HMI tags "Process_Value"
   "DB602_PV_Tank_Tank{0}_Temp_PV_Conf_ActV_ModulNo" : Int = PLC DB602_PV_Tank.Tank[0].Temp.PV_Conf_ActV.ModulNo AT %DB602.DBW32, 1 s
      on ChangeValue: SetBit("DB702_Tank_Value.Write")
   "DB602_PV_Tank_Tank{0}_Temp_PV_Conf_ActV_Address" : Int = PLC DB602_PV_Tank.Tank[0].Temp.PV_Conf_ActV.Address AT %DB602.DBW34, 1 s
      on ChangeValue: SetBit("DB702_Tank_Value.Write")
   "DB602_PV_Tank_Tank{0}_Temp_PV_Conf_ActV_OffsetSignal" : Int = PLC DB602_PV_Tank.Tank[0].Temp.PV_Conf_ActV.OffsetSignal AT %DB602.DBW36, 1 s
      on ChangeValue: SetBit("DB702_Tank_Value.Write")
   "DB602_PV_Tank_Tank{0}_Temp_PV_Conf_ActV_Multiplier" : Real = PLC DB602_PV_Tank.Tank[0].Temp.PV_Conf_ActV.Multiplier AT %DB602.DBD38, 1 s
      on ChangeValue: SetBit("DB702_Tank_Value.Write")
   "DB602_PV_Tank_Tank{0}_Temp_PV_Conf_ActV_MinValueSensor" : Real = PLC DB602_PV_Tank.Tank[0].Temp.PV_Conf_ActV.MinValueSensor AT %DB602.DBD42, 1 s
      on ChangeValue: SetBit("DB702_Tank_Value.Write")
   "DB602_PV_Tank_Tank{0}_Temp_PV_Conf_ActV_MaxValueSensor" : Real = PLC DB602_PV_Tank.Tank[0].Temp.PV_Conf_ActV.MaxValueSensor AT %DB602.DBD46, 1 s
      on ChangeValue: SetBit("DB702_Tank_Value.Write")
   "DB602_PV_Tank_Tank{0}_Temp_PV_Conf_ActV_MaxSignalResolution" : Real = PLC DB602_PV_Tank.Tank[0].Temp.PV_Conf_ActV.MaxSignalResolution AT %DB602.DBD50, 1 s
      on ChangeValue: SetBit("DB702_Tank_Value.Write")
   "DB602_PV_Tank_Tank{0}_Temp_PV_ActV_Value" : Real = PLC DB602_PV_Tank.Tank[0].Temp.PV_ActV.Value AT %DB602.DBD26, 1 s
      on ChangeValue: SetBit("DB702_Tank_Value.Write")
   "DB602_PV_Tank_Tank{0}_Level_PV_ActV_Value" : Real = PLC DB602_PV_Tank.Tank[0].Level.PV_ActV.Value AT %DB602.DBD74, 1 s
      on ChangeValue: SetBit("DB702_Tank_Value.Write")
   "DB602_PV_Tank_Tank{0}_Level_PV_Conf_ActV_ModulNo" : Int = PLC DB602_PV_Tank.Tank[0].Level.PV_Conf_ActV.ModulNo AT %DB602.DBW80, 1 s
      on ChangeValue: SetBit("DB702_Tank_Value.Write")
   "DB602_PV_Tank_Tank{0}_Level_PV_Conf_ActV_Address" : Int = PLC DB602_PV_Tank.Tank[0].Level.PV_Conf_ActV.Address AT %DB602.DBW82, 1 s
      on ChangeValue: SetBit("DB702_Tank_Value.Write")
   "DB602_PV_Tank_Tank{0}_Level_PV_Conf_ActV_OffsetSignal" : Int = PLC DB602_PV_Tank.Tank[0].Level.PV_Conf_ActV.OffsetSignal AT %DB602.DBW84, 1 s
      on ChangeValue: SetBit("DB702_Tank_Value.Write")
   "DB602_PV_Tank_Tank{0}_Level_PV_Conf_ActV_Multiplier" : Real = PLC DB602_PV_Tank.Tank[0].Level.PV_Conf_ActV.Multiplier AT %DB602.DBD86, 1 s
      on ChangeValue: SetBit("DB702_Tank_Value.Write")
   "DB602_PV_Tank_Tank{0}_Level_PV_Conf_ActV_MinValueSensor" : Real = PLC DB602_PV_Tank.Tank[0].Level.PV_Conf_ActV.MinValueSensor AT %DB602.DBD90, 1 s
      on ChangeValue: SetBit("DB702_Tank_Value.Write")
   "DB602_PV_Tank_Tank{0}_Level_PV_Conf_ActV_MaxValueSensor" : Real = PLC DB602_PV_Tank.Tank[0].Level.PV_Conf_ActV.MaxValueSensor AT %DB602.DBD94, 1 s
      on ChangeValue: SetBit("DB702_Tank_Value.Write")
   "DB602_PV_Tank_Tank{0}_Level_PV_Conf_ActV_MaxSignalResolution" : Real = PLC DB602_PV_Tank.Tank[0].Level.PV_Conf_ActV.MaxSignalResolution AT %DB602.DBD98, 1 s
      on ChangeValue: SetBit("DB702_Tank_Value.Write")
   "DB602_PV_Tank_Tank{0}_Nucleation_PV_Conf_ActV_ModulNo" : Int = PLC DB602_PV_Tank.Tank[0].Nucleation.PV_Conf_ActV.ModulNo AT %DB602.DBW176, 1 s
      on ChangeValue: SetBit("DB702_Tank_Value.Write")
   "DB602_PV_Tank_Tank{0}_Nucleation_PV_Conf_ActV_Address" : Int = PLC DB602_PV_Tank.Tank[0].Nucleation.PV_Conf_ActV.Address AT %DB602.DBW178, 1 s
      on ChangeValue: SetBit("DB702_Tank_Value.Write")
   "DB602_PV_Tank_Tank{0}_Nucleation_PV_Conf_ActV_OffsetSignal" : Int = PLC DB602_PV_Tank.Tank[0].Nucleation.PV_Conf_ActV.OffsetSignal AT %DB602.DBW180, 1 s
      on ChangeValue: SetBit("DB702_Tank_Value.Write")
   "DB602_PV_Tank_Tank{0}_Nucleation_PV_Conf_ActV_Multiplier" : Real = PLC DB602_PV_Tank.Tank[0].Nucleation.PV_Conf_ActV.Multiplier AT %DB602.DBD182, 1 s
      on ChangeValue: SetBit("DB702_Tank_Value.Write")
   "DB602_PV_Tank_Tank{0}_Nucleation_PV_Conf_ActV_MinValueSensor" : Real = PLC DB602_PV_Tank.Tank[0].Nucleation.PV_Conf_ActV.MinValueSensor AT %DB602.DBD186, 1 s
      on ChangeValue: SetBit("DB702_Tank_Value.Write")
   "DB602_PV_Tank_Tank{0}_Nucleation_PV_Conf_ActV_MaxValueSensor" : Real = PLC DB602_PV_Tank.Tank[0].Nucleation.PV_Conf_ActV.MaxValueSensor AT %DB602.DBD190, 1 s
      on ChangeValue: SetBit("DB702_Tank_Value.Write")
   "DB602_PV_Tank_Tank{0}_Nucleation_PV_Conf_ActV_MaxSignalResolution" : Real = PLC DB602_PV_Tank.Tank[0].Nucleation.PV_Conf_ActV.MaxSignalResolution AT %DB602.DBD194, 1 s
      on ChangeValue: SetBit("DB702_Tank_Value.Write")
   "DB602_PV_Tank_Tank{0}_Nucleation_PV_ActV_Value" : Real = PLC DB602_PV_Tank.Tank[0].Nucleation.PV_ActV.Value AT %DB602.DBD170, 1 s
      on ChangeValue: SetBit("DB702_Tank_Value.Write")
   "DB702_Tank_Value_Read" : Bool = PLC DB702_Tank_Value.Read AT %DB702.DBX4.0, 1 s
   "DB608_PV_Metering_Metering{0}_Flow_PV_Conf_ActV_Address" : Int = PLC DB608_PV_Metering.Metering[0].Flow.PV_Conf_ActV.Address AT %DB608.DBW34, 1 s
      on ChangeValue: SetBit("DB608_PV_Metering_Write")
   "DB608_PV_Metering_Metering{0}_Flow_PV_ActV_Value" : Real = PLC DB608_PV_Metering.Metering[0].Flow.PV_ActV.Value AT %DB608.DBD26, 1 s
      on ChangeValue: SetBit("DB608_PV_Metering_Write")
   "DB608_PV_Metering_Metering{0}_Pressure_PV_Conf_ActV_ModulNo" : Int = PLC DB608_PV_Metering.Metering[0].Pressure.PV_Conf_ActV.ModulNo AT %DB608.DBW80, 1 s
      on ChangeValue: SetBit("DB608_PV_Metering_Write")
   "DB608_PV_Metering_Metering{0}_Pressure_PV_Conf_ActV_Address" : Int = PLC DB608_PV_Metering.Metering[0].Pressure.PV_Conf_ActV.Address AT %DB608.DBW82, 1 s
      on ChangeValue: SetBit("DB608_PV_Metering_Write")
   "DB608_PV_Metering_Metering{0}_Pressure_PV_Conf_ActV_OffsetSignal" : Int = PLC DB608_PV_Metering.Metering[0].Pressure.PV_Conf_ActV.OffsetSignal AT %DB608.DBW84, 1 s
      on ChangeValue: SetBit("DB608_PV_Metering_Write")
   "DB608_PV_Metering_Metering{0}_Pressure_PV_Conf_ActV_Multiplier" : Real = PLC DB608_PV_Metering.Metering[0].Pressure.PV_Conf_ActV.Multiplier AT %DB608.DBD86, 1 s
      on ChangeValue: SetBit("DB608_PV_Metering_Write")
   "DB608_PV_Metering_Metering{0}_Pressure_PV_Conf_ActV_MinValueSensor" : Real = PLC DB608_PV_Metering.Metering[0].Pressure.PV_Conf_ActV.MinValueSensor AT %DB608.DBD90, 1 s
      on ChangeValue: SetBit("DB608_PV_Metering_Write")
   "DB608_PV_Metering_Metering{0}_Pressure_PV_Conf_ActV_MaxValueSensor" : Real = PLC DB608_PV_Metering.Metering[0].Pressure.PV_Conf_ActV.MaxValueSensor AT %DB608.DBD94, 1 s
      on ChangeValue: SetBit("DB608_PV_Metering_Write")
   "DB608_PV_Metering_Metering{0}_Pressure_PV_Conf_ActV_MaxSignalResolution" : Real = PLC DB608_PV_Metering.Metering[0].Pressure.PV_Conf_ActV.MaxSignalResolution AT %DB608.DBD98, 1 s
      on ChangeValue: SetBit("DB608_PV_Metering_Write")
   "DB608_PV_Metering_Metering{0}_Pressure_PV_ActV_Value" : Real = PLC DB608_PV_Metering.Metering[0].Pressure.PV_ActV.Value AT %DB608.DBD74, 1 s
      on ChangeValue: SetBit("DB608_PV_Metering_Write")
   "DB608_PV_Metering_Metering{0}_Temperature_PV_Conf_ActV_ModulNo" : Int = PLC DB608_PV_Metering.Metering[0].Temperature.PV_Conf_ActV.ModulNo AT %DB608.DBW128, 1 s
      on ChangeValue: SetBit("DB608_PV_Metering_Write")
   "DB608_PV_Metering_Metering{0}_Temperature_PV_Conf_ActV_Address" : Int = PLC DB608_PV_Metering.Metering[0].Temperature.PV_Conf_ActV.Address AT %DB608.DBW130, 1 s
      on ChangeValue: SetBit("DB608_PV_Metering_Write")
   "DB608_PV_Metering_Metering{0}_Temperature_PV_Conf_ActV_OffsetSignal" : Int = PLC DB608_PV_Metering.Metering[0].Temperature.PV_Conf_ActV.OffsetSignal AT %DB608.DBW132, 1 s
      on ChangeValue: SetBit("DB608_PV_Metering_Write")
   "DB608_PV_Metering_Metering{0}_Temperature_PV_Conf_ActV_Multiplier" : Real = PLC DB608_PV_Metering.Metering[0].Temperature.PV_Conf_ActV.Multiplier AT %DB608.DBD134, 1 s
      on ChangeValue: SetBit("DB608_PV_Metering_Write")
   "DB608_PV_Metering_Metering{0}_Temperature_PV_Conf_ActV_MinValueSensor" : Real = PLC DB608_PV_Metering.Metering[0].Temperature.PV_Conf_ActV.MinValueSensor AT %DB608.DBD138, 1 s
      on ChangeValue: SetBit("DB608_PV_Metering_Write")
   "DB608_PV_Metering_Metering{0}_Temperature_PV_Conf_ActV_MaxValueSensor" : Real = PLC DB608_PV_Metering.Metering[0].Temperature.PV_Conf_ActV.MaxValueSensor AT %DB608.DBD142, 1 s
      on ChangeValue: SetBit("DB608_PV_Metering_Write")
   "DB608_PV_Metering_Metering{0}_Temperature_PV_Conf_ActV_MaxSignalResolution" : Real = PLC DB608_PV_Metering.Metering[0].Temperature.PV_Conf_ActV.MaxSignalResolution AT %DB608.DBD146, 1 s
      on ChangeValue: SetBit("DB608_PV_Metering_Write")
   "DB608_PV_Metering_Metering{0}_Temperature_PV_ActV_Value" : Real = PLC DB608_PV_Metering.Metering[0].Temperature.PV_ActV.Value AT %DB608.DBD122, 1 s
      on ChangeValue: SetBit("DB608_PV_Metering_Write")
   "DB608_PV_Metering_Metering{0}_Pre_Pressure_PV_ActV_Value" : Real = PLC DB608_PV_Metering.Metering[0].Pre_Pressure.PV_ActV.Value AT %DB608.DBD170, 1 s
      on ChangeValue: SetBit("DB608_PV_Metering_Write")
   "DB608_PV_Metering_Metering{0}_Pre_Pressure_PV_Conf_ActV_ModulNo" : Int = PLC DB608_PV_Metering.Metering[0].Pre_Pressure.PV_Conf_ActV.ModulNo AT %DB608.DBW176, 1 s
      on ChangeValue: SetBit("DB608_PV_Metering_Write")
   "DB608_PV_Metering_Metering{0}_Pre_Pressure_PV_Conf_ActV_Address" : Int = PLC DB608_PV_Metering.Metering[0].Pre_Pressure.PV_Conf_ActV.Address AT %DB608.DBW178, 1 s
      on ChangeValue: SetBit("DB608_PV_Metering_Write")
   "DB608_PV_Metering_Metering{0}_Pre_Pressure_PV_Conf_ActV_OffsetSignal" : Int = PLC DB608_PV_Metering.Metering[0].Pre_Pressure.PV_Conf_ActV.OffsetSignal AT %DB608.DBW180, 1 s
      on ChangeValue: SetBit("DB608_PV_Metering_Write")
   "DB608_PV_Metering_Metering{0}_Pre_Pressure_PV_Conf_ActV_Multiplier" : Real = PLC DB608_PV_Metering.Metering[0].Pre_Pressure.PV_Conf_ActV.Multiplier AT %DB608.DBD182, 1 s
      on ChangeValue: SetBit("DB608_PV_Metering_Write")
   "DB608_PV_Metering_Metering{0}_Pre_Pressure_PV_Conf_ActV_MinValueSensor" : Real = PLC DB608_PV_Metering.Metering[0].Pre_Pressure.PV_Conf_ActV.MinValueSensor AT %DB608.DBD186, 1 s
      on ChangeValue: SetBit("DB608_PV_Metering_Write")
   "DB608_PV_Metering_Metering{0}_Pre_Pressure_PV_Conf_ActV_MaxValueSensor" : Real = PLC DB608_PV_Metering.Metering[0].Pre_Pressure.PV_Conf_ActV.MaxValueSensor AT %DB608.DBD190, 1 s
      on ChangeValue: SetBit("DB608_PV_Metering_Write")
   "DB608_PV_Metering_Metering{0}_Pre_Pressure_PV_Conf_ActV_MaxSignalResolution" : Real = PLC DB608_PV_Metering.Metering[0].Pre_Pressure.PV_Conf_ActV.MaxSignalResolution AT %DB608.DBD194, 1 s
      on ChangeValue: SetBit("DB608_PV_Metering_Write")
   "DB608_PV_Metering_HeatexchangerHP{0}_PV_ActV_Value" : Real = PLC DB608_PV_Metering.HeatexchangerHP[0].PV_ActV.Value AT %DB608.DBD3146, 1 s
      on ChangeValue: SetBit("DB608_PV_Metering_Write")
   "DB608_PV_Metering_HeatexchangerHP{0}_PV_Conf_ActV_ModulNo" : Int = PLC DB608_PV_Metering.HeatexchangerHP[0].PV_Conf_ActV.ModulNo AT %DB608.DBW3152, 1 s
      on ChangeValue: SetBit("DB608_PV_Metering_Write")
   "DB608_PV_Metering_HeatexchangerHP{0}_PV_Conf_ActV_Address" : Int = PLC DB608_PV_Metering.HeatexchangerHP[0].PV_Conf_ActV.Address AT %DB608.DBW3154, 1 s
      on ChangeValue: SetBit("DB608_PV_Metering_Write")
   "DB608_PV_Metering_HeatexchangerHP{0}_PV_Conf_ActV_OffsetSignal" : Int = PLC DB608_PV_Metering.HeatexchangerHP[0].PV_Conf_ActV.OffsetSignal AT %DB608.DBW3156, 1 s
      on ChangeValue: SetBit("DB608_PV_Metering_Write")
   "DB608_PV_Metering_HeatexchangerHP{0}_PV_Conf_ActV_Multiplier" : Real = PLC DB608_PV_Metering.HeatexchangerHP[0].PV_Conf_ActV.Multiplier AT %DB608.DBD3158, 1 s
      on ChangeValue: SetBit("DB608_PV_Metering_Write")
   "DB608_PV_Metering_HeatexchangerHP{0}_PV_Conf_ActV_MinValueSensor" : Real = PLC DB608_PV_Metering.HeatexchangerHP[0].PV_Conf_ActV.MinValueSensor AT %DB608.DBD3162, 1 s
      on ChangeValue: SetBit("DB608_PV_Metering_Write")
   "DB608_PV_Metering_HeatexchangerHP{0}_PV_Conf_ActV_MaxValueSensor" : Real = PLC DB608_PV_Metering.HeatexchangerHP[0].PV_Conf_ActV.MaxValueSensor AT %DB608.DBD3166, 1 s
      on ChangeValue: SetBit("DB608_PV_Metering_Write")
   "DB608_PV_Metering_HeatexchangerHP{0}_PV_Conf_ActV_MaxSignalResolution" : Real = PLC DB608_PV_Metering.HeatexchangerHP[0].PV_Conf_ActV.MaxSignalResolution AT %DB608.DBD3170, 1 s
      on ChangeValue: SetBit("DB608_PV_Metering_Write")
   "DB604_PV_Mixinghead_Mixinghead{0}_Inerting_PV_Conf_ActV_ModulNo" : Int = PLC DB604_PV_Mixinghead.Mixinghead[0].Inerting.PV_Conf_ActV.ModulNo AT %DB604.DBW704, 1 s
      on ChangeValue: SetBit("DB704_MH_Value_Write")
   "DB604_PV_Mixinghead_Mixinghead{0}_Inerting_PV_Conf_ActV_Address" : Int = PLC DB604_PV_Mixinghead.Mixinghead[0].Inerting.PV_Conf_ActV.Address AT %DB604.DBW706, 1 s
      on ChangeValue: SetBit("DB704_MH_Value_Write")
   "DB604_PV_Mixinghead_Mixinghead{0}_Inerting_PV_Conf_ActV_OffsetSignal" : Int = PLC DB604_PV_Mixinghead.Mixinghead[0].Inerting.PV_Conf_ActV.OffsetSignal AT %DB604.DBW708, 1 s
      on ChangeValue: SetBit("DB704_MH_Value_Write")
   "DB604_PV_Mixinghead_Mixinghead{0}_Inerting_PV_Conf_ActV_Multiplier" : Real = PLC DB604_PV_Mixinghead.Mixinghead[0].Inerting.PV_Conf_ActV.Multiplier AT %DB604.DBD710, 1 s
      on ChangeValue: SetBit("DB704_MH_Value_Write")
   "DB604_PV_Mixinghead_Mixinghead{0}_Inerting_PV_Conf_ActV_MinValueSensor" : Real = PLC DB604_PV_Mixinghead.Mixinghead[0].Inerting.PV_Conf_ActV.MinValueSensor AT %DB604.DBD714, 1 s
      on ChangeValue: SetBit("DB704_MH_Value_Write")
   "DB604_PV_Mixinghead_Mixinghead{0}_Inerting_PV_Conf_ActV_MaxValueSensor" : Real = PLC DB604_PV_Mixinghead.Mixinghead[0].Inerting.PV_Conf_ActV.MaxValueSensor AT %DB604.DBD718, 1 s
      on ChangeValue: SetBit("DB704_MH_Value_Write")
   "DB604_PV_Mixinghead_Mixinghead{0}_Inerting_PV_Conf_ActV_MaxSignalResolution" : Real = PLC DB604_PV_Mixinghead.Mixinghead[0].Inerting.PV_Conf_ActV.MaxSignalResolution AT %DB604.DBD722, 1 s
      on ChangeValue: SetBit("DB704_MH_Value_Write")
   "DB604_PV_Mixinghead_Mixinghead{0}_Inerting_PV_ActV_Value" : Real = PLC DB604_PV_Mixinghead.Mixinghead[0].Inerting.PV_ActV.Value AT %DB604.DBD698, 1 s
      on ChangeValue: SetBit("DB704_MH_Value_Write")
   "DB604_PV_Mixinghead_Mixinghead{0}_Pressure_Connection{1}_PV_Conf_ActV_ModulNo" : Int = PLC DB604_PV_Mixinghead.Mixinghead[0].Pressure_Connection[1].PV_Conf_ActV.ModulNo AT %DB604.DBW32, 1 s
      on ChangeValue: SetBit("DB704_MH_Value_Write")
   "DB604_PV_Mixinghead_Mixinghead{0}_Pressure_Connection{1}_PV_Conf_ActV_Address" : Int = PLC DB604_PV_Mixinghead.Mixinghead[0].Pressure_Connection[1].PV_Conf_ActV.Address AT %DB604.DBW34, 1 s
      on ChangeValue: SetBit("DB704_MH_Value_Write")
   "DB604_PV_Mixinghead_Mixinghead{0}_Pressure_Connection{1}_PV_Conf_ActV_OffsetSignal" : Int = PLC DB604_PV_Mixinghead.Mixinghead[0].Pressure_Connection[1].PV_Conf_ActV.OffsetSignal AT %DB604.DBW36, 1 s
      on ChangeValue: SetBit("DB704_MH_Value_Write")
   "DB604_PV_Mixinghead_Mixinghead{0}_Pressure_Connection{1}_PV_Conf_ActV_Multiplier" : Real = PLC DB604_PV_Mixinghead.Mixinghead[0].Pressure_Connection[1].PV_Conf_ActV.Multiplier AT %DB604.DBD38, 1 s
      on ChangeValue: SetBit("DB704_MH_Value_Write")
   "DB604_PV_Mixinghead_Mixinghead{0}_Pressure_Connection{1}_PV_Conf_ActV_MinValueSensor" : Real = PLC DB604_PV_Mixinghead.Mixinghead[0].Pressure_Connection[1].PV_Conf_ActV.MinValueSensor AT %DB604.DBD42, 1 s
      on ChangeValue: SetBit("DB704_MH_Value_Write")
   "DB604_PV_Mixinghead_Mixinghead{0}_Pressure_Connection{1}_PV_Conf_ActV_MaxValueSensor" : Real = PLC DB604_PV_Mixinghead.Mixinghead[0].Pressure_Connection[1].PV_Conf_ActV.MaxValueSensor AT %DB604.DBD46, 1 s
      on ChangeValue: SetBit("DB704_MH_Value_Write")
   "DB604_PV_Mixinghead_Mixinghead{0}_Pressure_Connection{1}_PV_Conf_ActV_MaxSignalResolution" : Real = PLC DB604_PV_Mixinghead.Mixinghead[0].Pressure_Connection[1].PV_Conf_ActV.MaxSignalResolution AT %DB604.DBD50, 1 s
      on ChangeValue: SetBit("DB704_MH_Value_Write")
   "DB604_PV_Mixinghead_Mixinghead{0}_Pressure_Connection{2}_PV_Conf_ActV_ModulNo" : Int = PLC DB604_PV_Mixinghead.Mixinghead[0].Pressure_Connection[2].PV_Conf_ActV.ModulNo AT %DB604.DBW80, 1 s
      on ChangeValue: SetBit("DB704_MH_Value_Write")
   "DB604_PV_Mixinghead_Mixinghead{0}_Pressure_Connection{2}_PV_Conf_ActV_Address" : Int = PLC DB604_PV_Mixinghead.Mixinghead[0].Pressure_Connection[2].PV_Conf_ActV.Address AT %DB604.DBW82, 1 s
      on ChangeValue: SetBit("DB704_MH_Value_Write")
   "DB604_PV_Mixinghead_Mixinghead{0}_Pressure_Connection{2}_PV_Conf_ActV_OffsetSignal" : Int = PLC DB604_PV_Mixinghead.Mixinghead[0].Pressure_Connection[2].PV_Conf_ActV.OffsetSignal AT %DB604.DBW84, 1 s
      on ChangeValue: SetBit("DB704_MH_Value_Write")
   "DB604_PV_Mixinghead_Mixinghead{0}_Pressure_Connection{2}_PV_Conf_ActV_Multiplier" : Real = PLC DB604_PV_Mixinghead.Mixinghead[0].Pressure_Connection[2].PV_Conf_ActV.Multiplier AT %DB604.DBD86, 1 s
      on ChangeValue: SetBit("DB704_MH_Value_Write")
   "DB604_PV_Mixinghead_Mixinghead{0}_Pressure_Connection{2}_PV_Conf_ActV_MinValueSensor" : Real = PLC DB604_PV_Mixinghead.Mixinghead[0].Pressure_Connection[2].PV_Conf_ActV.MinValueSensor AT %DB604.DBD90, 1 s
      on ChangeValue: SetBit("DB704_MH_Value_Write")
   "DB604_PV_Mixinghead_Mixinghead{0}_Pressure_Connection{2}_PV_Conf_ActV_MaxValueSensor" : Real = PLC DB604_PV_Mixinghead.Mixinghead[0].Pressure_Connection[2].PV_Conf_ActV.MaxValueSensor AT %DB604.DBD94, 1 s
      on ChangeValue: SetBit("DB704_MH_Value_Write")
   "DB604_PV_Mixinghead_Mixinghead{0}_Pressure_Connection{2}_PV_Conf_ActV_MaxSignalResolution" : Real = PLC DB604_PV_Mixinghead.Mixinghead[0].Pressure_Connection[2].PV_Conf_ActV.MaxSignalResolution AT %DB604.DBD98, 1 s
      on ChangeValue: SetBit("DB704_MH_Value_Write")
   "DB604_PV_Mixinghead_Mixinghead{0}_Pressure_Connection{3}_PV_Conf_ActV_ModulNo" : Int = PLC DB604_PV_Mixinghead.Mixinghead[0].Pressure_Connection[3].PV_Conf_ActV.ModulNo AT %DB604.DBW128, 1 s
      on ChangeValue: SetBit("DB704_MH_Value_Write")
   "DB604_PV_Mixinghead_Mixinghead{0}_Pressure_Connection{3}_PV_Conf_ActV_Address" : Int = PLC DB604_PV_Mixinghead.Mixinghead[0].Pressure_Connection[3].PV_Conf_ActV.Address AT %DB604.DBW130, 1 s
      on ChangeValue: SetBit("DB704_MH_Value_Write")
   "DB604_PV_Mixinghead_Mixinghead{0}_Pressure_Connection{3}_PV_Conf_ActV_OffsetSignal" : Int = PLC DB604_PV_Mixinghead.Mixinghead[0].Pressure_Connection[3].PV_Conf_ActV.OffsetSignal AT %DB604.DBW132, 1 s
      on ChangeValue: SetBit("DB704_MH_Value_Write")
   "DB604_PV_Mixinghead_Mixinghead{0}_Pressure_Connection{3}_PV_Conf_ActV_Multiplier" : Real = PLC DB604_PV_Mixinghead.Mixinghead[0].Pressure_Connection[3].PV_Conf_ActV.Multiplier AT %DB604.DBD134, 1 s
      on ChangeValue: SetBit("DB704_MH_Value_Write")
   "DB604_PV_Mixinghead_Mixinghead{0}_Pressure_Connection{3}_PV_Conf_ActV_MinValueSensor" : Real = PLC DB604_PV_Mixinghead.Mixinghead[0].Pressure_Connection[3].PV_Conf_ActV.MinValueSensor AT %DB604.DBD138, 1 s
      on ChangeValue: SetBit("DB704_MH_Value_Write")
   "DB604_PV_Mixinghead_Mixinghead{0}_Pressure_Connection{3}_PV_Conf_ActV_MaxValueSensor" : Real = PLC DB604_PV_Mixinghead.Mixinghead[0].Pressure_Connection[3].PV_Conf_ActV.MaxValueSensor AT %DB604.DBD142, 1 s
      on ChangeValue: SetBit("DB704_MH_Value_Write")
   "DB604_PV_Mixinghead_Mixinghead{0}_Pressure_Connection{3}_PV_Conf_ActV_MaxSignalResolution" : Real = PLC DB604_PV_Mixinghead.Mixinghead[0].Pressure_Connection[3].PV_Conf_ActV.MaxSignalResolution AT %DB604.DBD146, 1 s
      on ChangeValue: SetBit("DB704_MH_Value_Write")
   "DB604_PV_Mixinghead_Mixinghead{0}_Pressure_Connection{4}_PV_Conf_ActV_ModulNo" : Int = PLC DB604_PV_Mixinghead.Mixinghead[0].Pressure_Connection[4].PV_Conf_ActV.ModulNo AT %DB604.DBW176, 1 s
      on ChangeValue: SetBit("DB704_MH_Value_Write")
   "DB604_PV_Mixinghead_Mixinghead{0}_Pressure_Connection{4}_PV_Conf_ActV_Address" : Int = PLC DB604_PV_Mixinghead.Mixinghead[0].Pressure_Connection[4].PV_Conf_ActV.Address AT %DB604.DBW178, 1 s
      on ChangeValue: SetBit("DB704_MH_Value_Write")
   "DB604_PV_Mixinghead_Mixinghead{0}_Pressure_Connection{4}_PV_Conf_ActV_OffsetSignal" : Int = PLC DB604_PV_Mixinghead.Mixinghead[0].Pressure_Connection[4].PV_Conf_ActV.OffsetSignal AT %DB604.DBW180, 1 s
      on ChangeValue: SetBit("DB704_MH_Value_Write")
   "DB604_PV_Mixinghead_Mixinghead{0}_Pressure_Connection{4}_PV_Conf_ActV_Multiplier" : Real = PLC DB604_PV_Mixinghead.Mixinghead[0].Pressure_Connection[4].PV_Conf_ActV.Multiplier AT %DB604.DBD182, 1 s
      on ChangeValue: SetBit("DB704_MH_Value_Write")
   "DB604_PV_Mixinghead_Mixinghead{0}_Pressure_Connection{4}_PV_Conf_ActV_MinValueSensor" : Real = PLC DB604_PV_Mixinghead.Mixinghead[0].Pressure_Connection[4].PV_Conf_ActV.MinValueSensor AT %DB604.DBD186, 1 s
      on ChangeValue: SetBit("DB704_MH_Value_Write")
   "DB604_PV_Mixinghead_Mixinghead{0}_Pressure_Connection{4}_PV_Conf_ActV_MaxValueSensor" : Real = PLC DB604_PV_Mixinghead.Mixinghead[0].Pressure_Connection[4].PV_Conf_ActV.MaxValueSensor AT %DB604.DBD190, 1 s
      on ChangeValue: SetBit("DB704_MH_Value_Write")
   "DB604_PV_Mixinghead_Mixinghead{0}_Pressure_Connection{4}_PV_Conf_ActV_MaxSignalResolution" : Real = PLC DB604_PV_Mixinghead.Mixinghead[0].Pressure_Connection[4].PV_Conf_ActV.MaxSignalResolution AT %DB604.DBD194, 1 s
      on ChangeValue: SetBit("DB704_MH_Value_Write")
   "DB604_PV_Mixinghead_Mixinghead{0}_Pressure_Connection{5}_PV_Conf_ActV_ModulNo" : Int = PLC DB604_PV_Mixinghead.Mixinghead[0].Pressure_Connection[5].PV_Conf_ActV.ModulNo AT %DB604.DBW224, 1 s
      on ChangeValue: SetBit("DB704_MH_Value_Write")
   "DB604_PV_Mixinghead_Mixinghead{0}_Pressure_Connection{5}_PV_Conf_ActV_Address" : Int = PLC DB604_PV_Mixinghead.Mixinghead[0].Pressure_Connection[5].PV_Conf_ActV.Address AT %DB604.DBW226, 1 s
      on ChangeValue: SetBit("DB704_MH_Value_Write")
   "DB604_PV_Mixinghead_Mixinghead{0}_Pressure_Connection{5}_PV_Conf_ActV_OffsetSignal" : Int = PLC DB604_PV_Mixinghead.Mixinghead[0].Pressure_Connection[5].PV_Conf_ActV.OffsetSignal AT %DB604.DBW228, 1 s
      on ChangeValue: SetBit("DB704_MH_Value_Write")
   "DB604_PV_Mixinghead_Mixinghead{0}_Pressure_Connection{5}_PV_Conf_ActV_Multiplier" : Real = PLC DB604_PV_Mixinghead.Mixinghead[0].Pressure_Connection[5].PV_Conf_ActV.Multiplier AT %DB604.DBD230, 1 s
      on ChangeValue: SetBit("DB704_MH_Value_Write")
   "DB604_PV_Mixinghead_Mixinghead{0}_Pressure_Connection{5}_PV_Conf_ActV_MinValueSensor" : Real = PLC DB604_PV_Mixinghead.Mixinghead[0].Pressure_Connection[5].PV_Conf_ActV.MinValueSensor AT %DB604.DBD234, 1 s
      on ChangeValue: SetBit("DB704_MH_Value_Write")
   "DB604_PV_Mixinghead_Mixinghead{0}_Pressure_Connection{5}_PV_Conf_ActV_MaxValueSensor" : Real = PLC DB604_PV_Mixinghead.Mixinghead[0].Pressure_Connection[5].PV_Conf_ActV.MaxValueSensor AT %DB604.DBD238, 1 s
      on ChangeValue: SetBit("DB704_MH_Value_Write")
   "DB604_PV_Mixinghead_Mixinghead{0}_Pressure_Connection{5}_PV_Conf_ActV_MaxSignalResolution" : Real = PLC DB604_PV_Mixinghead.Mixinghead[0].Pressure_Connection[5].PV_Conf_ActV.MaxSignalResolution AT %DB604.DBD242, 1 s
      on ChangeValue: SetBit("DB704_MH_Value_Write")
   "DB604_PV_Mixinghead_Mixinghead{0}_Pressure_Connection{6}_PV_Conf_ActV_ModulNo" : Int = PLC DB604_PV_Mixinghead.Mixinghead[0].Pressure_Connection[6].PV_Conf_ActV.ModulNo AT %DB604.DBW272, 1 s
      on ChangeValue: SetBit("DB704_MH_Value_Write")
   "DB604_PV_Mixinghead_Mixinghead{0}_Pressure_Connection{6}_PV_Conf_ActV_Address" : Int = PLC DB604_PV_Mixinghead.Mixinghead[0].Pressure_Connection[6].PV_Conf_ActV.Address AT %DB604.DBW274, 1 s
      on ChangeValue: SetBit("DB704_MH_Value_Write")
   "DB604_PV_Mixinghead_Mixinghead{0}_Pressure_Connection{6}_PV_Conf_ActV_OffsetSignal" : Int = PLC DB604_PV_Mixinghead.Mixinghead[0].Pressure_Connection[6].PV_Conf_ActV.OffsetSignal AT %DB604.DBW276, 1 s
      on ChangeValue: SetBit("DB704_MH_Value_Write")
   "DB604_PV_Mixinghead_Mixinghead{0}_Pressure_Connection{6}_PV_Conf_ActV_Multiplier" : Real = PLC DB604_PV_Mixinghead.Mixinghead[0].Pressure_Connection[6].PV_Conf_ActV.Multiplier AT %DB604.DBD278, 1 s
      on ChangeValue: SetBit("DB704_MH_Value_Write")
   "DB604_PV_Mixinghead_Mixinghead{0}_Pressure_Connection{6}_PV_Conf_ActV_MinValueSensor" : Real = PLC DB604_PV_Mixinghead.Mixinghead[0].Pressure_Connection[6].PV_Conf_ActV.MinValueSensor AT %DB604.DBD282, 1 s
      on ChangeValue: SetBit("DB704_MH_Value_Write")
   "DB604_PV_Mixinghead_Mixinghead{0}_Pressure_Connection{6}_PV_Conf_ActV_MaxValueSensor" : Real = PLC DB604_PV_Mixinghead.Mixinghead[0].Pressure_Connection[6].PV_Conf_ActV.MaxValueSensor AT %DB604.DBD286, 1 s
      on ChangeValue: SetBit("DB704_MH_Value_Write")
   "DB604_PV_Mixinghead_Mixinghead{0}_Pressure_Connection{6}_PV_Conf_ActV_MaxSignalResolution" : Real = PLC DB604_PV_Mixinghead.Mixinghead[0].Pressure_Connection[6].PV_Conf_ActV.MaxSignalResolution AT %DB604.DBD290, 1 s
      on ChangeValue: SetBit("DB704_MH_Value_Write")
   "DB604_PV_Mixinghead_Mixinghead{0}_Temperature_Connection{1}_PV_Conf_ActV_ModulNo" : Int = PLC DB604_PV_Mixinghead.Mixinghead[0].Temperature_Connection[1].PV_Conf_ActV.ModulNo AT %DB604.DBW320, 1 s
      on ChangeValue: SetBit("DB704_MH_Value_Write")
   "DB604_PV_Mixinghead_Mixinghead{0}_Temperature_Connection{1}_PV_Conf_ActV_Address" : Int = PLC DB604_PV_Mixinghead.Mixinghead[0].Temperature_Connection[1].PV_Conf_ActV.Address AT %DB604.DBW322, 1 s
      on ChangeValue: SetBit("DB704_MH_Value_Write")
   "DB604_PV_Mixinghead_Mixinghead{0}_Temperature_Connection{1}_PV_Conf_ActV_OffsetSignal" : Int = PLC DB604_PV_Mixinghead.Mixinghead[0].Temperature_Connection[1].PV_Conf_ActV.OffsetSignal AT %DB604.DBW324, 1 s
      on ChangeValue: SetBit("DB704_MH_Value_Write")
   "DB604_PV_Mixinghead_Mixinghead{0}_Temperature_Connection{1}_PV_Conf_ActV_Multiplier" : Real = PLC DB604_PV_Mixinghead.Mixinghead[0].Temperature_Connection[1].PV_Conf_ActV.Multiplier AT %DB604.DBD326, 1 s
      on ChangeValue: SetBit("DB704_MH_Value_Write")
   "DB604_PV_Mixinghead_Mixinghead{0}_Temperature_Connection{1}_PV_Conf_ActV_MinValueSensor" : Real = PLC DB604_PV_Mixinghead.Mixinghead[0].Temperature_Connection[1].PV_Conf_ActV.MinValueSensor AT %DB604.DBD330, 1 s
      on ChangeValue: SetBit("DB704_MH_Value_Write")
   "DB604_PV_Mixinghead_Mixinghead{0}_Temperature_Connection{1}_PV_Conf_ActV_MaxValueSensor" : Real = PLC DB604_PV_Mixinghead.Mixinghead[0].Temperature_Connection[1].PV_Conf_ActV.MaxValueSensor AT %DB604.DBD334, 1 s
      on ChangeValue: SetBit("DB704_MH_Value_Write")
   "DB604_PV_Mixinghead_Mixinghead{0}_Temperature_Connection{1}_PV_Conf_ActV_MaxSignalResolution" : Real = PLC DB604_PV_Mixinghead.Mixinghead[0].Temperature_Connection[1].PV_Conf_ActV.MaxSignalResolution AT %DB604.DBD338, 1 s
      on ChangeValue: SetBit("DB704_MH_Value_Write")
   "DB604_PV_Mixinghead_Mixinghead{0}_Temperature_Connection{2}_PV_Conf_ActV_ModulNo" : Int = PLC DB604_PV_Mixinghead.Mixinghead[0].Temperature_Connection[2].PV_Conf_ActV.ModulNo AT %DB604.DBW368, 1 s
      on ChangeValue: SetBit("DB704_MH_Value_Write")
   "DB604_PV_Mixinghead_Mixinghead{0}_Temperature_Connection{2}_PV_Conf_ActV_Address" : Int = PLC DB604_PV_Mixinghead.Mixinghead[0].Temperature_Connection[2].PV_Conf_ActV.Address AT %DB604.DBW370, 1 s
      on ChangeValue: SetBit("DB704_MH_Value_Write")
   "DB604_PV_Mixinghead_Mixinghead{0}_Temperature_Connection{2}_PV_Conf_ActV_OffsetSignal" : Int = PLC DB604_PV_Mixinghead.Mixinghead[0].Temperature_Connection[2].PV_Conf_ActV.OffsetSignal AT %DB604.DBW372, 1 s
      on ChangeValue: SetBit("DB704_MH_Value_Write")
   "DB604_PV_Mixinghead_Mixinghead{0}_Temperature_Connection{2}_PV_Conf_ActV_Multiplier" : Real = PLC DB604_PV_Mixinghead.Mixinghead[0].Temperature_Connection[2].PV_Conf_ActV.Multiplier AT %DB604.DBD374, 1 s
      on ChangeValue: SetBit("DB704_MH_Value_Write")
   "DB604_PV_Mixinghead_Mixinghead{0}_Temperature_Connection{2}_PV_Conf_ActV_MinValueSensor" : Real = PLC DB604_PV_Mixinghead.Mixinghead[0].Temperature_Connection[2].PV_Conf_ActV.MinValueSensor AT %DB604.DBD378, 1 s